        .INPUT_xSyncroPhotocell_1   // M403.P115B1.Synchro photocell / start count
        .PH_x.0   // Load
        .PH_x.1   // Load Upstream
        .PH_x.10   // Unload Upstream
        .PH_x.11   // End load Downstream
        .PH_x.12   // Unload Downstream
        .PH_x.13   // End unload Upstream
        .PH_x.14   // End unload Downstream
        .PH_x.15   // End unload
        .PH_x.16   // Unload Unpack (n caps)
        .PH_x.17   // End unload Unpack (n caps)
        .PH_x.18   // Unload Unpack (n caps) Upstream
        .PH_x.19   // End unload Unpack (n caps) Upstream
        .PH_x.2   // Load Downstream
        .PH_x.20   // Unload Unpack (n caps) Downstream
        .PH_x.21   // End unload Unpack (n caps) Downstream
        .PH_x.22   // Load reentry
        .PH_x.23   // End load reentry
        .PH_x.24   // Unload reentry
        .PH_x.25   // End unload reentry
        .PH_x.26   // Load Unpack (n caps)
        .PH_x.27   // End load Unpack (n caps)
        .PH_x.28   // Load Unpack (n caps) Upstream
        .PH_x.29   // End load Unpack (n caps) Upstream
        .PH_x.3   // Wait rotation done
        .PH_x.30   // Load Unpack (n caps) Downstream
        .PH_x.31   // End load Unpack (n caps) Downstream
        .PH_x.4   // Rotation ended
        .PH_x.7   // End load
        .PH_x.8   // Unload
        .PH_x.9   // End load Upstream
   M316_ALM : MAC_Conveyor_ALM;
        .rgdFaultCode_M[0]   // Drive fault code M1
        .rgdFaultCode_M[1]   // Drive fault code M2
        .rgxStoppingFault[0].0   // Z402.M316-M1.Positioning error
        .rgxStoppingFault[0].1   // Z402.M316-M1.Phase in progress with rotator not in low position
        .rgxStoppingFault_M[0].0   // Z402.M316-M1.Protection motor rotation
        .rgxStoppingFault_M[0].1   // Z402.M316-M1.Drive error
        .rgxStoppingFault_M[0].2   // Z402.M316-M1.Drive feedback error
        .rgxStoppingFault_M[0].3   // Z402.M316-M1.Local safety switch
        .rgxStoppingFault_M[0].4   // Z402.M316-M1.Motor thermal probe
        .rgxStoppingFault_M[0].5   // Z402.M316-M1.Braking resistor anomaly
        .rgxStoppingFault_M[0].6   // Z402.M316-M1.Drive not ready
        .rgxWarning[0].0   // Z402.M316.Plate not synchronized
        .rgxWarning[0].1   // Z402.M316.Positioning error
   M316_Data : UDT_Convoy_SL;
   M316_dLastRotationA_ID : DINT; {access Read Only}
   M316_HMR : MAC_Conveyor_HMR := (xIdPlatePresence := 1, dState1 := 1, dState2 := 1, dStateSensor1 := 1, dStateSensor2 := 1, dStateSensor3 := 1, dStateSensor4 := 1);
        .dErrorCode1   // Error code M1
        .rgxMan.0   // Run M1
        .rgxMan.1   // Reverse M1
        .rgxMan.2   // Run M2
        .rgxMan.3   // Reverse M2
        .rgxMan.4   // Run both
        .rgxMan.5   // Reverse both
        .dErrorCode2   // Error code M2
        .xSensorPresence1   // M403.P115B1.Synchro photocell / start count {x|x|x|x|O}
        .xSensorPresence2   // M403.P115B2.Synchro photocell / start count {x|x|x|x|O}
   M316_HMW : MAC_Conveyor_HMW;
        .dParam_1_cmm   // Positioning offset 1 [mm] {mm/100|mm|-50|+50|M}
        .dParam_2_cmm   // Positioning offset 2 [mm] {mm/100|mm|-50|+50|M}
        .rgxMan.0   // Run M1
        .rgxMan.1   // Reverse M1
        .rgxMan.2   // Run M2
        .rgxMan.3   // Reverse M2
        .rgxMan.4   // Run both
        .rgxMan.5   // Reverse both
   M316_M1_DR : AXIS_CIP_DRIVE; {access Read Only}
   M316_M1_DR_IN_MAJ : MOTION_INSTRUCTION := (FLAGS := 570425344, DN := 1); {access None}
   M316_M1_DR_IN_MAM : MOTION_INSTRUCTION := (FLAGS := 704643072, DN := 1, PC := 1); {access None}
   M316_M1_DR_IN_MAR : MOTION_INSTRUCTION := (FLAGS := 167772160, PC := 1); {access None}
   M316_M1_DR_IN_MAS : MOTION_INSTRUCTION := (FLAGS := -1442840576, EN := 1, DN := 1, PC := 1); {access None}
   M316_M1_DR_IN_MCD : MOTION_INSTRUCTION := (FLAGS := 570425344, DN := 1); {access None}
   M316_M1_DR_IN_MRP : MOTION_INSTRUCTION := (FLAGS := 536870912, DN := 1, STATUS := 2, STATE := 3); {access None}
   M316_M1_DR_MAFR : MOTION_INSTRUCTION := (FLAGS := 301989888, ER := 1, ERR := 11); {access None}
   M316_M1_DR_MDR : MOTION_INSTRUCTION := (FLAGS := -1845493760, EN := 1, ER := 1, ERR := 11); {access None}
   M316_M1_DR_MSF : MOTION_INSTRUCTION := (FLAGS := 570425344, DN := 1, STATUS := 2, STATE := 1); {access None}
   M316_M1_DR_MSO : MOTION_INSTRUCTION := (FLAGS := -1610612736, EN := 1, DN := 1, STATE := 1); {access None}
   M316_M1_DR_OUT_MAJ : MOTION_INSTRUCTION := (FLAGS := 570425344, DN := 1); {access None}
   M316_M1_DR_OUT_MAM : MOTION_INSTRUCTION := (FLAGS := 704643072, DN := 1, PC := 1); {access None}
   M316_M1_DR_OUT_MAR : MOTION_INSTRUCTION := (FLAGS := 671088640, DN := 1, PC := 1, STATE := 1); {access None}
   M316_M1_DR_OUT_MAS : MOTION_INSTRUCTION := (FLAGS := -1442840576, EN := 1, DN := 1, PC := 1); {access None}
   M316_M1_DR_OUT_MCD : MOTION_INSTRUCTION := (FLAGS := 570425344, DN := 1); {access None}
   M316_M1_DR_OUT_MRP : MOTION_INSTRUCTION := (FLAGS := 536870912, DN := 1, STATUS := 2, STATE := 3); {access None}
   M316_SpaceConv_Utilities : SpaceConv_Utilities := (CONST_dSyncMode := 1, CONST_dSyncroPhWindow_cmm := 450000, CONST_dConveyorLength_cmm := 800000, CONST_dConveyorWidth_cmm := 400000, CONST_dPresetFeedbackTime_ms := 500, CONST_rAcceleration_ms2 := 1.2, CONST_rDeceleration_ms2 := 1.2, CONF_MD1_dScan_ms := 20, CONF_MD2_MD3_dPrstPos_cmm := -390000, CONF_MD4_MD6_dLength_cmm := 365800, CONF_MD7_dOffset_cmm := 50000, ST_dStopLoadForseen_cmm := 620000, ST_dRealSpeed_mm_min := 90000, ST_rStepAdvancementH := 3000.0, ST_rStepAdvancementT := 3000.0, O_xPlateSynchronized := 1, O_dCountFeedbackTime_ms := 500, O_dPresetLoadUnload_cmm := -126300);
   M316_TON_Synchro_timeout : TIMER; {access Read Only}
   M316_xOS_SentToCullet : BOOL; {access Read Only}
   M316_xPlateCullet : BOOL; {access Read Only}
   M316_xSendCulletReqActive : BOOL; {access Read Only}
   M316_xSensorTimeout : BOOL; {access Read Only}
   M316A : MAC_Rotator := (ST_xCleaningConditionOK := 1, ST_xConditionOKStopCycle := 1, ST_xEnableControlError := 1, INPUT_rRotatorPosition_cdeg := 26999.898, INPUT_xConditionToDescent := 1, INPUT_xLowPosition := 1, INPUT_xLocalSafetySwitchRotation := 1, INPUT_xProtectionMotorLifting := 1, INPUT_xProtectionMotorRotation := 1, tmON_DelayFrameUP.PRE := 100, tmON_DelayRotatorInRun.PRE := 300, tmOF_DriveEnable.PRE := 20000, tmOF_DriveEnable.ACC := 20000, tmON_FeedbackTimeOutLifting.PRE := 1000, tmON_FeedbackTimeOutRotation.PRE := 1000, tmON_FramePosError.PRE := 2500, tmON_RotatePosError.PRE := 10000, tmON_RotatePosError.ACC := 2040, tmON_RotatePosError.EN := 1, tmON_RotatePosError.TT := 1, tmON_PresetEncoder.PRE := 3000, tmON_DelayBrakeON.PRE := 200); {access None}
        .OUTPUT_xDescent   // P253KA4.Descent frame
        .PH_x.0   // Rise frame
        .PH_x.12   // Counterclockwise rotation
        .PH_x.4   // Descent frame
        .PH_x.8   // Clockwise totation
        .OUTPUT_xRise   // P253KA3.Lifting frame
        .INPUT_xLowPosition   // P56KA2.Frame to low position
        .INPUT_xFeedbackLifting   // P56KM1/2.Feedback lifting chassis
        .INPUT_xHighPosition   // P56KA1.Frame to high position
        .INPUT_xProtectionMotorLifting   // P56QM1.Protection lifting frame
   M316A_ALM : MAC_Rotator_ALM;
        .rgxStoppingFault_M[0].0   // Z402.M316A.Protection motor rotation
        .rgxStoppingFault_M[0].1   // Z402.M316A.Drive Error
        .rgxStoppingFault_M[0].11   // Z402.M316A.Frame lifting position error
        .rgxStoppingFault_M[0].2   // Z402.M316A.Drive feedback error
        .rgxStoppingFault_M[0].20   // Z402.M316A.Drive not ready
        .rgxStoppingFault_M[0].3   // Z402.M316A.Rotation position error
        .rgxStoppingFault_M[0].8   // Z402.M316A.Protection lifting frame
        .rgxStoppingFault_M[0].9   // Z402.M316A.Feedback lifting chassis
   M316A_Data : UDT_Convoy_SL;
   M316A_HMR : MAC_Rotator_HMR := (xLowPosition := 1, dState := 1, dActualAngle_cdeg := 27000);
        .rgxMan.0   // Rise
        .rgxMan.1   // Descent
        .rgxMan.10   // Clockwise rotation jog
        .rgxMan.11   // Counter Clockwise rotation jog
        .rgxMan.14   // Enable brake release
        .rgxMan.15   // Disable brake release
        .rgxMan.8   // Clockwise rotation
        .rgxMan.9   // Counter Clockwise rotation
   M316A_HMW : MAC_Rotator_HMW := (xPresetEnc := 1, dLowSpeed_deg_s := 40, dLowRamp_deg_s2 := 50, dHighSpeed_deg_s := 50, dHighRamp_deg_s2 := 60, dJogSpeed_deg_s := 12);
        .rgxMan.0   // Rise
        .rgxMan.1   // Descent
        .rgxMan.10   // Clockwise rotation jog
        .rgxMan.11   // Counterclockwise rotation jog
        .rgxMan.14   // Enable brake release
        .rgxMan.15   // Disable brake release
        .rgxMan.8   // Clockwise rotation
        .rgxMan.9   // Counterclockwise rotation
   M316A_M1_DR : AXIS_CIP_DRIVE; {access Read Only}
   M316A_M1_DR_IN_MAJ : MOTION_INSTRUCTION := (FLAGS := 570425344, DN := 1); {access None}
   M316A_M1_DR_IN_MAM : MOTION_INSTRUCTION := (FLAGS := 704643072, DN := 1, PC := 1); {access None}
   M316A_M1_DR_IN_MAS : MOTION_INSTRUCTION := (FLAGS := -1442840576, EN := 1, DN := 1, PC := 1); {access None}
   M316A_M1_DR_MAFR : MOTION_INSTRUCTION := (FLAGS := 301989888, ER := 1, ERR := 11); {access None}
   M316A_M1_DR_MAH : MOTION_INSTRUCTION := (FLAGS := 671088640, DN := 1, PC := 1, STATE := 17); {access None}
   M316A_M1_DR_MSF : MOTION_INSTRUCTION := (FLAGS := -1610612736, EN := 1, DN := 1, STATUS := 2, STATE := 1); {access None}
   M316A_M1_DR_MSO : MOTION_INSTRUCTION := (FLAGS := 536870912, DN := 1, STATE := 1); {access None}
   M316A_M1_DR_OUT_MAJ : MOTION_INSTRUCTION := (FLAGS := 570425344, DN := 1); {access None}
   M316A_M1_DR_OUT_MAM : MOTION_INSTRUCTION := (FLAGS := 704643072, DN := 1, PC := 1); {access None}
   M316A_M1_DR_OUT_MAS : MOTION_INSTRUCTION := (FLAGS := -1442840576, EN := 1, DN := 1, PC := 1); {access None}
   M316A_MAM_IP_TOFF : TIMER; {access Read Only}
   M316A_rLastPosition : REAL; {access Read Only}
   M316A_TmON1 : TIMER; {access Read Only}
   M316M317_OffsetBaricentre_cmm : DINT; {access Read Only}
   M317 : MAC_Conveyor_Single := (ST_xCleaningConditionOK := 1, ST_xPlatePresence := 1, ST_xConditionOKStopCycle := 1, ST_xOutputEnable := 1, ST_xIdPlatePresence := 1, ST_xWaitStopNextMachine := 1, ST_xEnableControlError := 1, ST_xPlateSynchronized := 1, ST_xSafetyMovement := 1, OSR_xSynchroPhotocellTail := 1, INPUT_xSquaringPhotocell_4 := 1, INPUT_xLowPositionSquaring_1 := 1, INPUT_xHighPositionPopup_1 := 1, INPUT_xHighPositionPopup_2 := 1, INPUT_xDriveReady_M1 := 1, INPUT_xLocalSafetySwitch_M1 := 1, INPUT_xMotorThermalProbe_M1 := 1, INPUT_xProtectionMotor_M1 := 1, INPUT_xDriveReady_M2 := 1, INPUT_xLocalSafetySwitch_M2 := 1, INPUT_xMotorThermalProbe_M2 := 1, INPUT_xProtectionMotor_M2 := 1, INPUT_xDriveFeedback_M3 := 1, INPUT_xDriveReady_M3 := 1, INPUT_xLocalSafetySwitch_M3 := 1, INPUT_xMotorThermalProbe_M3 := 1, INPUT_xProtectionMotor_M3 := 1, INPUT_xDriveReady_M4 := 1, INPUT_xLocalSafetySwitch_M4 := 1, INPUT_xMotorThermalProbe_M4 := 1, INPUT_xProtectionMotor_M4 := 1, INPUT_xProtectionLiftingFrame_1 := 1, INPUT_xProtectionLiftingFrame_2 := 1, INPUT_xFeedbackVentilation_1 := 1, INPUT_xFeedbackVentilation_2 := 1, OUTPUT_xDriveEnable_M1 := 1, OUTPUT_xDriveEnable_M2 := 1, OUTPUT_xDriveEnable_M3 := 1, OUTPUT_xDriveEnable_M4 := 1, OUTPUT_xFunCommand_1 := 1, OUTPUT_xFunCommand_2 := 1, AUX_dPresetStopLoad_cmm := 372333, AUX_dPresetStopUnload_cmm := 441667, AUX_dAccSpace_cmm := 41667, AUX_dDecSpace_cmm := 41667, AUX_dReqSpeed_mm_min := 60000, AUX_dAbsPosTarget_M3_cmm := 195500, AUX_dAbsPosTarget_M4_cmm := 195500, AUX_dQtaLites := 1, tmON_FeedbackTimeOut_M1.PRE := 2000, tmOF_DriveEnable_M1.PRE := 30000, tmOF_DriveEnable_M1.ACC := 540, tmOF_DriveEnable_M1.TT := 1, tmOF_DriveEnable_M1.DN := 1, tmOF_PowerSaving_M1.EN := 1, tmOF_PowerSaving_M1.DN := 1, tmON_FeedbackTimeOut_M2.PRE := 2000, tmOF_DriveEnable_M2.PRE := 30000, tmOF_DriveEnable_M2.ACC := 540, tmOF_DriveEnable_M2.TT := 1,
        tmOF_DriveEnable_M2.DN := 1, tmON_FeedbackTimeOut_M3.PRE := 2000, tmOF_DriveEnable_M3.PRE := 30000, tmOF_DriveEnable_M3.ACC := 540, tmOF_DriveEnable_M3.TT := 1, tmOF_DriveEnable_M3.DN := 1, tmON_FeedbackTimeOut_M4.PRE := 2000, tmOF_DriveEnable_M4.PRE := 30000, tmOF_DriveEnable_M4.ACC := 540, tmOF_DriveEnable_M4.TT := 1, tmOF_DriveEnable_M4.DN := 1, tmON_AuxFunction1.PRE := 5000, tmON_AuxFunction1.EN := 1, tmON_AuxFunction1.DN := 1, tmON_AuxFunction2.PRE := 2200, tmON_AuxFunction3.PRE := 2200, tmON_AuxFunction4.PRE := 15000, tmON_AuxFunction5.PRE := 3000, tmON_AuxFunction6.PRE := 15000, tmON_AuxFunction7.PRE := 3600000, tmON_AuxFunction8.PRE := 40000, tmON_AuxFunction9.PRE := 20000, TmON[0].PRE := 3000, TmON[1].PRE := 1000, TmON[1].ACC := 1019, TmON[2].PRE := 5000, TmON[6].PRE := 5000, TmON[6].EN := 1, TmON[6].DN := 1, TmON[11].PRE := 2000, TmON[12].PRE := 2000, TmON[13].PRE := 2000, TmON[14].PRE := 2000, tmOF_MCD_M1.ACC := 20, tmOF_MCD_M2.ACC := 20, tmOF_MCD_M3.ACC := 20, tmOF_MCD_M4.ACC := 20); {access None}
        .INPUT_xSquaringPhotocell_1   // P406B1.Squaring frontal photocell - Right
        .INPUT_xMotorThermalProbe_M2   // M2.P404BT2.Motor thermal probe
        .INPUT_xLowPositionPopup_1   // P63KA2.M5.Low position popup
        .INPUT_xLowPositionSquaring_1   // P405SQ2.Low position squaring
        .INPUT_xMotorThermalProbe_M1   // M1.P404BT1.Motor thermal probe
        .INPUT_xHighPositionPopup_1   // P63KA1.M5.High position popup
        .INPUT_xSquaringPhotocell_2   // P406B2.Squaring frontal photocell - Left
        .INPUT_xHighPositionPopup_2   // P64KA1.M6.High position popup
        .PH_x.0   // Load (from M316)
        .PH_x.10   // Load (from M419)
        .PH_x.11   // End load (from M419)
        .PH_x.12   // Unload (to M316)
        .PH_x.13   // End unload (to M316)
        .PH_x.15   // End unload (to M419)
        .PH_x.16   // Rise popup
        .PH_x.19   // End rise popup
        .PH_x.20   // Descent popup
        .PH_x.23   // End descent popup
        .PH_x.24   // Reset counter position
        .PH_x.26   // Lateral positioning (M3-M4)
        .PH_x.27   // End lateral positioning (M3-M4)
        .PH_x.28   // Lateral squaring
        .PH_x.29   // End lateral squaring
        .PH_x.30   // Lateral traction recovery (M3-M4)
        .PH_x.31   // End lateral traction recovery (M3-M4)
        .PH_x.4   // Frontal squaring (run fwd + rise squaring)
        .PH_x.5   // End frontal sqauring
        .PH_x.7   // End load (from M316)
        .PH_x.8   // Unload (to M419)
        .INPUT_xMotorThermalProbe_M3   // M3.P405BT3.Motor thermal probe
        .INPUT_xLowPositionPopup_2   // P64KA2.M6.Low position popup
        .INPUT_xSquaringPhotocell_3   // P405B1.Squaring lateral photocell - Right
        .INPUT_xHighPositionSquaring_1   // P405SQ1.High position squaring
        .INPUT_xSquaringPhotocell_4   // P405B2.Squaring lateral photocell - Left
        .INPUT_xHighPositionSquaring_2   // P405SQ11.High position squaring
        .ST_xAux1   // Ready to unload on backward conveyor
        .INPUT_xLowPositionSquaring_2   // P405SQ12.Low position squaring
   M317_ALM : MAC_Conveyor_ALM;
        .rgxWarning[0].10   // Z402.M317-M2.Plate not synchronized
        .rgdFaultCode_M[0]   // Drive fault code M1
        .rgdFaultCode_M[1]   // Drive fault code M2
        .rgxStoppingFault[0].0   // Z402.M317-M1.Positioning error
        .rgxStoppingFault[0].1   // Z402.M317-M1.Plate not synchronized
        .rgxStoppingFault[0].10   // Z402.M317-M2.Error position frontal squaring
        .rgxStoppingFault[0].11   // Z402.M317-M2.Timeout frontal squaring
        .rgxStoppingFault[0].12   // Z402.M317-M2.Lugs position sensors fault
        .rgxStoppingFault[0].13   // Z402.M317. Timeout movement popup 1
        .rgxStoppingFault[0].14   // Z402.M317. Timeout movement popup 2
        .rgxStoppingFault[0].16   // Z402.M317-M3.Positioning error
        .rgxStoppingFault[0].18   // Z402.M317-M3.Error position popup
        .rgxStoppingFault[0].19   // Z402.M317-M3.Error position lateral squaring
        .rgxStoppingFault[0].2   // Z402.M317-M1.Error position frontal squaring
        .rgxStoppingFault[0].20   // Z402.M317-M3.Timeout lateral squaring
        .rgxStoppingFault[0].21   // Z402.M317.Protection lifting popup 1
        .rgxStoppingFault[0].22   // Z402.M317.Protection lifting popup 2
        .rgxStoppingFault[0].3   // Z402.M317-M1.Timeout frontal squaring
        .rgxStoppingFault[0].4   // Z402.M317-M1.Lugs position sensors fault
        .rgxStoppingFault[0].5   // Z402.M317. Popup 1 position error
        .rgxStoppingFault[0].6   // Z402.M317. Popup 2 position error
        .rgxStoppingFault[0].8   // Z402.M317-M2.Positioning error
        .rgxStoppingFault[0].9   // Z402.M317-M2.Plate not synchronized
        .rgxStoppingFault_M[0].0   // Z402.M317-M1.P59AZ1.Protection motor rotation
        .rgxStoppingFault_M[0].1   // Z402.M317-M1.P59AZ1.Drive error
        .rgxStoppingFault_M[0].10   // Z402.M317-M2.P59AZ1.Drive feedback error
        .rgxStoppingFault_M[0].11   // Z402.M317-M2.P59AZ1.Local safety switch
        .rgxStoppingFault_M[0].12   // Z402.M317-M2.P405BT2.Motor thermal probe
        .rgxStoppingFault_M[0].13   // Z402.M317-M2.P59AZ1.Braking resistor anomaly
        .rgxStoppingFault_M[0].14   // Z402.M317-M2.Drive not ready
        .rgxStoppingFault_M[0].16   // Z402.M317-M3.P61AZ1.Protection motor rotation
        .rgxStoppingFault_M[0].17   // Z402.M317-M3.P61AZ1.Drive error
        .rgxStoppingFault_M[0].18   // Z402.M317-M3.P61AZ1.Drive feedback error
        .rgxStoppingFault_M[0].19   // Z402.M317-M3.P61AZ1.Local safety switch
        .rgxStoppingFault_M[0].2   // Z402.M317-M1.P59AZ1.Drive feedback error
        .rgxStoppingFault_M[0].20   // Z402.M317-M3.P404BT1.Motor thermal probe
        .rgxStoppingFault_M[0].21   // Z402.M317-M3.Drive not ready
        .rgxStoppingFault_M[0].3   // Z402.M317-M1.P59AZ1.Local safety switch
        .rgxStoppingFault_M[0].4   // Z402.M317-M1.P405BT1.Motor thermal probe
        .rgxStoppingFault_M[0].5   // Z402.M317-M1.P59AZ1.Braking resistor anomaly
        .rgxStoppingFault_M[0].6   // Z402.M317-M1.Drive not ready
        .rgxStoppingFault_M[0].8   // Z402.M317-M2.P59AZ1.Protection motor rotation
        .rgxStoppingFault_M[0].9   // Z402.M317-M2.P59AZ1.Drive error
        .rgxWarning[0].0   // Z402.M317-M1.Plate not synchronized
        .rgxWarning[0].1   // Z402.M317-M1.Positioning error
        .rgxWarning[0].11   // Z402.M317-M2.Positioning error
        .rgxWarning[0].21   // Z402.M317-M3.Lateal positioning error
        .rgxWarning[0].25   // Z402.M317.Timeout frontal squaring
        .rgxWarning[0].26   // Z402.M317.Timeout lateral squaring
   M317_AlmTimer1 : TIMER; {access Read Only}
   M317_AlmTimer2 : TIMER; {access Read Only}
   M317_Data : UDT_Convoy_SL;
        .rgtCap[0].rgxRequest.0   // Frontal squaring request
        .rgtCap[0].rgxRequest.1   // Lateral squaring request
        .rgtCap[0].rgxRequest.2   // Y adjust position request
        .rgtCap[0].rgxRequest.3   // Y measure request
        .rgtCap[0].rgxDone.0   // Frontal squaring done
        .rgtCap[0].rgxDone.1   // Lateral squaring done
        .rgtCap[0].rgxDone.2   // Y adjust position done
        .rgtCap[0].rgxDone.3   // Y measure done
   M317_dSlowingSquaringQuote : DINT; {access Read Only}
   M317_dTractionRecovery_M3 : DINT; {access Read Only}
   M317_dTractionRecovery_M4 : DINT; {access Read Only}
   M317_HMR : MAC_Conveyor_HMR := (xSensorPresence4 := 1, xHighPositionPopup1 := 1, xHighPositionPopup2 := 1, xLowPositionSquaring1 := 1, xLowPositionSquaring2 := 1, xIdPlatePresence := 1, dState1 := 1, dState2 := 1, dState3 := 1, dState4 := 1, dStateSensor1 := 1, dStateSensor2 := 1, dStateSensor3 := 1, dStateSensor4 := 1, dStateSensor5 := 1, dStateSensor6 := 1);
        .xSensorPresence5   // P115/3.Start count photocell {x|x|x|x|O}
        .xHighPositionPopup2   // P64KA1.M6.High position popup {x|x|x|x|O}
        .dErrorCode1   // Error code M1
        .xHighPositionPopup1   // P63KA1.M5.High position popup {x|x|x|x|O}
        .rgxMan.0   // Run M1
        .rgxMan.1   // Reverse M1
        .rgxMan.10   // Rise popup 1
        .rgxMan.11   // Descent popup 1
        .rgxMan.12   // Rise popup 2
        .rgxMan.13   // Descent popup 2
        .rgxMan.14   // Rise all popups
        .rgxMan.15   // Descent all popups
        .rgxMan.16   // Rise frontal squaring 1
        .rgxMan.17   // Descent frontal squaring 1
        .rgxMan.18   // Rise frontal squaring 2
        .rgxMan.19   // Descent frontal squaring 2
        .rgxMan.2   // Run M2
        .rgxMan.20   // Rise all frontal squaring
        .rgxMan.21   // Descent all frontal squaring
        .rgxMan.3   // Reverse M2
        .rgxMan.4   // Run M3
        .rgxMan.5   // Reverse M3
        .rgxMan.6   // Run M4
        .rgxMan.7   // Reverse M4
        .dState3   // State M3 (1=No anomaly; 3=Run; 4=Reverse; 7=Anomaly)
        .xHighPositionSquaring1   // P405SQ1.High position frontal squaring M1 {x|x|x|x|O}
        .dErrorCode2   // Error code M2
        .xSensorPresence6   // P115/4.Start count photocell {x|x|x|x|O}
        .xSensorPresence4   // P404B1.SlowDown photocell frontal squaring left {x|x|x|x|O}
        .xLowPositionPopup1   // P63KA2.M5.Low position popup {x|x|x|x|O}
        .xHighPositionSquaring2   // P405SQ11.High position frontal squaring M2 {x|x|x|x|O}
        .dState2   // State M2 (1=No anomaly; 3=Run; 4=Reverse; 7=Anomaly)
        .dErrorCode4   // Error code M4
        .xSensorPresence3   // P404B1.SlowDown photocell frontal squaring right {x|x|x|x|O}
        .dState1   // State M1 (1=No anomaly; 3=Run; 4=Reverse; 7=Anomaly)
        .dState4   // State M4 (1=No anomaly; 3=Run; 4=Reverse; 7=Anomaly)
        .xLowPositionSquaring2   // P405SQ12.Low position frontal squaring M2 {x|x|x|x|O}
        .xLowPositionSquaring1   // P405SQ2.Low position frontal squaring M1 {x|x|x|x|O}
        .xLowPositionPopup2   // P64KA2.M6.Low position popup {x|x|x|x|O}
        .xSensorPresence1   // P405B1.SlowDown photocell lateral squaring right {x|x|x|x|O}
        .dErrorCode3   // Error code M3
        .xSensorPresence2   // P405B2.SlowDown photocell lateral squaring left {x|x|x|x|O}
   M317_HMW : MAC_Conveyor_HMW := (dParam_3_cmm := 4000, dParam_5_ms := 3000, dParam_6_ms := 4000, dParam_7_ms := 2200, dParam_8_ms := 5000);
        .dParam_4_cmm   // Lateral squaring space {mm/100|mm|0|500|M}
        .dParam_1_cmm   // Positioning offset 1 {mm/100|mm|-50|+50|M}
        .dParam_3_cmm   // Frontal squaring space {mm/100|mm|0|500|M}
        .dParam_6_ms   // Squaring frontal time 2 {ms|s|0|5|M}
        .dParam_2_cmm   // Positioning offset 2 {mm/100|mm|-50|+50|M}
        .dParam_8_ms   // Squaring lateral time 2 {ms|s|0|5|M}
        .rgxMan.0   // Run M1
        .rgxMan.1   // Reverse M1
        .rgxMan.10   // Rise popup 2
        .rgxMan.11   // Descent popup 2
        .rgxMan.12   // Rise all popups
        .rgxMan.13   // Descent all popups
        .rgxMan.14   // Run both (M1-2)
        .rgxMan.15   // Reverse both (M1-2)
        .rgxMan.16   // Rise frontal squaring 1
        .rgxMan.17   // Descent frontal squaring 1
        .rgxMan.18   // Rise frontal squaring 2
        .rgxMan.19   // Descent frontal squaring 2
        .rgxMan.2   // Run M2
        .rgxMan.20   // Rise all frontal squaring
        .rgxMan.21   // Descent all frontal squaring
        .rgxMan.3   // Reverse M2
        .rgxMan.4   // Run M3
        .rgxMan.5   // Reverse M3
        .rgxMan.6   // Run M4
        .rgxMan.7   // Reverse M4
        .rgxMan.8   // Rise popup 1
        .rgxMan.9   // Descent popup 1
        .dParam_7_ms   // Squaring lateral time 1 {ms|s|0|5|M}
        .dParam_5_ms   // Squaring frontal time 1 {ms|s|0|5|M}
   M317_M1_DR_IN_MAJ : MOTION_INSTRUCTION := (FLAGS := 570425344, DN := 1); {access None}
   M317_M1_DR_IN_MAM : MOTION_INSTRUCTION := (FLAGS := 33554432); {access None}
   M317_M1_DR_IN_MAR : MOTION_INSTRUCTION := (FLAGS := 33554432); {access None}
   M317_M1_DR_IN_MAS : MOTION_INSTRUCTION := (FLAGS := -1442840576, EN := 1, DN := 1, PC := 1); {access None}
   M317_M1_DR_IN_MCD : MOTION_INSTRUCTION := (FLAGS := 570425344, DN := 1); {access None}
   M317_M1_DR_IN_MRP : MOTION_INSTRUCTION := (FLAGS := 33554432); {access None}
   M317_M1_DR_MAFR : MOTION_INSTRUCTION := (FLAGS := 301989888, ER := 1, ERR := 11); {access None}
   M317_M1_DR_MDR : MOTION_INSTRUCTION := (FLAGS := -1845493760, EN := 1, ER := 1, ERR := 11); {access None}
   M317_M1_DR_MSF : MOTION_INSTRUCTION := (FLAGS := 570425344, DN := 1, STATUS := 2, STATE := 1); {access None}
   M317_M1_DR_MSO : MOTION_INSTRUCTION := (FLAGS := -1610612736, EN := 1, DN := 1, STATE := 1); {access None}
   M317_M1_DR_OUT_MAJ : MOTION_INSTRUCTION := (FLAGS := 570425344, DN := 1); {access None}
   M317_M1_DR_OUT_MAM : MOTION_INSTRUCTION := (FLAGS := 33554432); {access None}
   M317_M1_DR_OUT_MAR : MOTION_INSTRUCTION := (FLAGS := 33554432); {access None}
   M317_M1_DR_OUT_MAS : MOTION_INSTRUCTION := (FLAGS := -1442840576, EN := 1, DN := 1, PC := 1); {access None}
   M317_M1_DR_OUT_MCD : MOTION_INSTRUCTION := (FLAGS := 570425344, DN := 1); {access None}
   M317_M1_DR_OUT_MRP : MOTION_INSTRUCTION := (FLAGS := 33554432); {access None}
   M317_M1_DR_R1 : AXIS_CIP_DRIVE; {access Read Only}
   M317_M2_AUX_ReqSpeed_mm_min : DINT; {access Read Only}
   M317_M2_ChangeSpeed : BOOL; {access Read Only}
   M317_M2_DR_IN_MAJ : MOTION_INSTRUCTION := (FLAGS := 570425344, DN := 1); {access None}
   M317_M2_DR_IN_MAM : MOTION_INSTRUCTION := (FLAGS := 33554432); {access None}
   M317_M2_DR_IN_MAR : MOTION_INSTRUCTION := (FLAGS := 33554432); {access None}
   M317_M2_DR_IN_MAS : MOTION_INSTRUCTION := (FLAGS := 704643072, DN := 1, PC := 1); {access None}
   M317_M2_DR_IN_MCD : MOTION_INSTRUCTION := (FLAGS := 301989888, ER := 1, ERR := 23); {access None}
   M317_M2_DR_IN_MRP : MOTION_INSTRUCTION := (FLAGS := 536870912, DN := 1, STATUS := 2, STATE := 3); {access None}
   M317_M2_DR_MAFR : MOTION_INSTRUCTION := (FLAGS := 301989888, ER := 1, ERR := 11); {access None}
   M317_M2_DR_MDR : MOTION_INSTRUCTION := (FLAGS := -1845493760, EN := 1, ER := 1, ERR := 11); {access None}
   M317_M2_DR_MSF : MOTION_INSTRUCTION := (FLAGS := 570425344, DN := 1, STATUS := 2, STATE := 1); {access None}
   M317_M2_DR_MSO : MOTION_INSTRUCTION := (FLAGS := -1610612736, EN := 1, DN := 1, STATE := 1); {access None}
   M317_M2_DR_OUT_MAJ : MOTION_INSTRUCTION := (FLAGS := 570425344, DN := 1); {access None}
   M317_M2_DR_OUT_MAM : MOTION_INSTRUCTION := (FLAGS := 33554432); {access None}
   M317_M2_DR_OUT_MAR : MOTION_INSTRUCTION := (FLAGS := 33554432); {access None}
   M317_M2_DR_OUT_MAS : MOTION_INSTRUCTION := (FLAGS := 704643072, DN := 1, PC := 1); {access None}
   M317_M2_DR_OUT_MCD : MOTION_INSTRUCTION := (FLAGS := 301989888, ER := 1, ERR := 23); {access None}
   M317_M2_DR_OUT_MRP : MOTION_INSTRUCTION := (FLAGS := 536870912, DN := 1, STATUS := 2, STATE := 3); {access None}
   M317_M2_DR_R2 : AXIS_CIP_DRIVE; {access Read Only}
   M317_M2_ReqSpeed_mm_min : DINT; {access Read Only}
   M317_M3_AUX_ReqSpeed_mm_min : DINT; {access Read Only}
   M317_M3_ChangeSpeed : BOOL; {access Read Only}
   M317_M3_DR_IN_MAJ : MOTION_INSTRUCTION := (FLAGS := 570425344, DN := 1); {access None}
   M317_M3_DR_IN_MAM : MOTION_INSTRUCTION := (FLAGS := -1509949440, EN := 1, DN := 1, IP := 1); {access None}
   M317_M3_DR_IN_MAR : MOTION_INSTRUCTION := (FLAGS := 33554432); {access None}
   M317_M3_DR_IN_MAS : MOTION_INSTRUCTION := (FLAGS := 704643072, DN := 1, PC := 1); {access None}
   M317_M3_DR_IN_MCD : MOTION_INSTRUCTION := (FLAGS := 570425344, DN := 1); {access None}
   M317_M3_DR_IN_MRP : MOTION_INSTRUCTION := (FLAGS := 536870912, DN := 1, STATUS := 2, STATE := 3); {access None}
   M317_M3_DR_L : AXIS_CIP_DRIVE; {access Read Only}
   M317_M3_DR_MAFR : MOTION_INSTRUCTION := (FLAGS := 301989888, ER := 1, ERR := 11); {access None}
   M317_M3_DR_MDR : MOTION_INSTRUCTION := (FLAGS := -1845493760, EN := 1, ER := 1, ERR := 11); {access None}
   M317_M3_DR_MSF : MOTION_INSTRUCTION := (FLAGS := 570425344, DN := 1, STATUS := 2, STATE := 1); {access None}
   M317_M3_DR_MSO : MOTION_INSTRUCTION := (FLAGS := -1610612736, EN := 1, DN := 1, STATE := 1); {access None}
   M317_M3_DR_OUT_MAJ : MOTION_INSTRUCTION := (FLAGS := 570425344, DN := 1); {access None}
   M317_M3_DR_OUT_MAM : MOTION_INSTRUCTION := (FLAGS := -1509949440, EN := 1, DN := 1, IP := 1);
   M317_M3_DR_OUT_MAR : MOTION_INSTRUCTION := (FLAGS := 33554432); {access None}
   M317_M3_DR_OUT_MAS : MOTION_INSTRUCTION := (FLAGS := 704643072, DN := 1, PC := 1); {access None}
   M317_M3_DR_OUT_MCD : MOTION_INSTRUCTION := (FLAGS := 570425344, DN := 1); {access None}
   M317_M3_DR_OUT_MRP : MOTION_INSTRUCTION := (FLAGS := 536870912, DN := 1, STATUS := 2, STATE := 3); {access None}
   M317_M3_ReqSpeed_mm_min : DINT; {access Read Only}
   M317_M3_xOSR_LatSquarFtc : BOOL; {access Read Only}
   M317_SpaceConv_Utilities : SpaceConv_Utilities := (CONST_dSyncMode := 1, CONST_dSyncroPhWindow_cmm := 450000, CONST_dConveyorLength_cmm := 800000, CONST_dConveyorWidth_cmm := 400000, CONST_dPresetFeedbackTime_ms := 500, CONST_rAcceleration_ms2 := 1.2, CONST_rDeceleration_ms2 := 1.2, CONF_MD1_dScan_ms := 20, CONF_MD2_MD3_dPrstPos_cmm := -390000, CONF_MD4_MD6_dLength_cmm := 365800, CONF_MD7_dOffset_cmm := 50000, ST_dStopLoadForseen_cmm := 620000, ST_dRealSpeed_mm_min := 90000, ST_rStepAdvancementH := 3000.0, ST_rStepAdvancementT := 3000.0, O_xPlateSynchronized := 1, O_dCountFeedbackTime_ms := 500, O_dPresetLoadUnload_cmm := -126300);
   M317_TimerAlm3 : TIMER; {access Read Only}
   M317_TON_FrontSquarLeft_timeout : TIMER; {access Read Only}
   M317_TON_FrontSquarRight_timeout : TIMER; {access Read Only}
   M317_TON_LatSquarLeft_timeout : TIMER; {access Read Only}
   M317_TON_LatSquarRight_timeout : TIMER; {access Read Only}
   M317_TON_Load : TIMER; {access Read Only}
   M317_TON_Synchro_timeout : TIMER; {access Read Only}
   M317_xEnableTractionRecovering : BOOL; {access Read Only}
   M317_xFrontLeftTimeout : BOOL; {access Read Only}
   M317_xFrontRightTimeout : BOOL; {access Read Only}
   M317_xLateralTractionRecovered : BOOL; {access Read Only}
   M317_xLatLeftTimeout : BOOL; {access Read Only}
   M317_xLatRightTimeout : BOOL; {access Read Only}
   M317_xOS_PosReq : BOOL;
   M317_xPlateCullet : BOOL; {access Read Only}
   M317_xSendCulletReqActive : BOOL; {access Read Only}
   M317_xSensorTimeout : BOOL; {access Read Only}
   M350_M1_DR : AXIS_CIP_DRIVE; {access Read Only}
   M350_xReqStopPrevConvForPos : BOOL; {access Read Only}
   M350Popup : MAC_Popup_ZC; {access Read Only}
   M350Popup_ALM : MAC_Popup_ZC_ALM; {access Read Only}
        .rgxStoppingFault[0].0   // M350.Lifting position error
   M350Popup_DATA : UDT_ConvoyCap_ZC; {access Read Only}
   M350Popup_HMR : MAC_Popup_ZC_HMR := (xLowPosition := 1, rgdState := 1); {access Read Only}
        .rgxMan.0   // Rise popup {x|x|x|x|O}
        .rgxMan.1   // Lower popup {x|x|x|x|O}
   M350Popup_HMW : MAC_Popup_ZC_HMW := (dSingleCapOffset_cmm := 30000, dGlassPosFromStart_cmm := 15000, dGlassPosFromEnd_cmm := 15000, dConvoySidePosForCenterSheet := 1, dConvoyGapForCenterSheet := 50000, dSaturationSelection := 3);
        .rgxMan.0   // Rise popup {x|x|x|x|O}
        .rgxMan.1   // Lower popup {x|x|x|x|O}
   M350Popup_IN_MOTION : MAC_Popup_ZC_IN_MOTION; {access None}
   M350Popup_OUT_MOTION : MAC_Popup_ZC_OUT_MOTION; {access None}
   M350Popup_PlateFreeTimeout : TIMER := (PRE := 5000); {access Read Only}
   M350Popup_ReentryCap : UDT_ConvoyCap_ZC;
   M350Popup_SearchResultAfter : GP_TrackingSearchPlate_STC;
   M350Popup_SL_DATA : UDT_Convoy_SL; {access Read Only}
   M350Popup_xDrivePosEnable : BOOL; {access Read Only}
   M350Popup_xQualityComing : BOOL; {access Read Only}
   M351 : MAC_Conveyor;
        .INPUT_xMotorThermalProbe_M1   // M315A.M1.Q403BT3. Motor thermal probe
        .PH_x.0   // Load
        .PH_x.1   // Load Upstream
        .PH_x.10   // Unload Downstream
        .PH_x.13   // End unload Upstream
        .PH_x.14   // End unload Downstream
        .PH_x.15   // End unload
        .PH_x.16   // Unpack convoy
        .PH_x.17   // End unpack convoy
        .PH_x.18   // Unpack convoy Upstream
        .PH_x.19   // End unpack convoy Upstream
        .PH_x.2   // Load Downstream
        .PH_x.20   // Unpack convoy Downstream
        .PH_x.21   // End unpack convoy Downstream
        .PH_x.22   // Stop for unload on main line
        .PH_x.23   // End stop for unload on main line
        .PH_x.24   // Stop for unload on main line Upstream
        .PH_x.25   // End stop for unload on main line Upstream
        .PH_x.26   // Stop for unload on main line Downstream
        .PH_x.27   // End stop for unload on main line Downstream
        .PH_x.28   // Load reentry
        .PH_x.29   // End load reentry
        .PH_x.5   // End load Upstream
        .PH_x.6   // End load Downstream
        .PH_x.7   // End load
        .PH_x.8   // Unload
        .PH_x.9   // Unload Upstream
   M351_ALM : MAC_Conveyor_ALM;
        .rgdFaultCode_M[0]   // Drive fault code
        .rgxStoppingFault_M[0].0   // Z900.M351-M1.Protection motor rotation
        .rgxStoppingFault_M[0].1   // Z900.M351-M1.Drive error
        .rgxStoppingFault_M[0].2   // Z900.M351-M1.Drive feedback error
        .rgxStoppingFault_M[0].3   // Z900.M351-M1.Local safety switch
        .rgxStoppingFault_M[0].4   // Z900.M351.M1. Motor thermal probe
        .rgxStoppingFault_M[0].5   // Z900.M351-M1.Braking resistor anomaly
        .rgxStoppingFault_M[0].6   // Z900.M351-M1.Drive not ready
   M351_Data : UDT_Convoy_SL;
   M351_HMR : MAC_Conveyor_HMR := (xManualCommandEnabled := 1, dState4 := 1);
        .dErrorCode1   // Error code M1
        .rgxMan.0   // Run M1
        .rgxMan.1   // Reverse M1
        .rgxMan.2   // Run M2
        .rgxMan.3   // Reverse M2
        .rgxMan.4   // Run M3
        .rgxMan.5   // Reverse M3
        .dErrorCode2   // Error code M2 (NU)
        .dErrorCode3   // Error code M3 (NU)
   M351_HMW : MAC_Conveyor_HMW;
        .rgxMan.0   // Run M1
        .rgxMan.1   // Reverse M1
        .rgxMan.2   // Run M2
        .rgxMan.3   // Reverse M2
        .rgxMan.4   // Run M3
        .rgxMan.5   // Reverse M3
   M351_M1_DR : AXIS_CIP_DRIVE; {access Read Only}
   M351_M1_DR_IN_MAJ : MOTION_INSTRUCTION := (FLAGS := 570425344, DN := 1); {access None}
   M351_M1_DR_IN_MAM : MOTION_INSTRUCTION := (FLAGS := 33554432); {access None}
   M351_M1_DR_IN_MAR : MOTION_INSTRUCTION := (FLAGS := 33554432); {access None}
   M351_M1_DR_IN_MAS : MOTION_INSTRUCTION := (FLAGS := -1442840576, EN := 1, DN := 1, PC := 1); {access None}
   M351_M1_DR_IN_MCD : MOTION_INSTRUCTION := (FLAGS := 570425344, DN := 1); {access None}
   M351_M1_DR_IN_MRP : MOTION_INSTRUCTION := (FLAGS := 33554432); {access None}
   M351_M1_DR_MAFR : MOTION_INSTRUCTION := (FLAGS := 301989888, ER := 1, ERR := 11); {access None}
   M351_M1_DR_MDR : MOTION_INSTRUCTION := (FLAGS := -1845493760, EN := 1, ER := 1, ERR := 11); {access None}
   M351_M1_DR_MSF : MOTION_INSTRUCTION := (FLAGS := 536870912, DN := 1, STATUS := 2, STATE := 1); {access None}
   M351_M1_DR_MSO : MOTION_INSTRUCTION := (FLAGS := -1577058304, EN := 1, DN := 1, STATE := 1); {access None}
   M351_M1_DR_OUT_MAJ : MOTION_INSTRUCTION := (FLAGS := 570425344, DN := 1); {access None}
   M351_M1_DR_OUT_MAM : MOTION_INSTRUCTION := (FLAGS := 33554432); {access None}
   M351_M1_DR_OUT_MAR : MOTION_INSTRUCTION := (FLAGS := 33554432); {access None}
   M351_M1_DR_OUT_MAS : MOTION_INSTRUCTION := (FLAGS := -1442840576, EN := 1, DN := 1, PC := 1); {access None}
   M351_M1_DR_OUT_MCD : MOTION_INSTRUCTION := (FLAGS := 570425344, DN := 1); {access None}
   M351_M1_DR_OUT_MRP : MOTION_INSTRUCTION := (FLAGS := 33554432); {access None}
   M351_SpaceConv_Utilities : SpaceConv_Utilities := (CONST_dSyncMode := 1, CONST_dSyncroPhWindow_cmm := 200000, CONST_dConveyorLength_cmm := 500000, CONST_dConveyorWidth_cmm := 400000, CONST_dPresetFeedbackTime_ms := 500, CONST_rAcceleration_ms2 := 1.2, CONST_rDeceleration_ms2 := 1.2, CONF_MD1_dScan_ms := 20, CONF_MD4_MD6_dLength_cmm := 360000, CONF_MD7_dOffset_cmm := 50000, ST_xLastModLoadBkw := 1, ST_dStopLoadForseen_cmm := 495370, ST_dRealSpeed_mm_min := 40000, ST_rStepAdvancementH := 1333.3334, ST_rStepAdvancementT := 1333.3334, O_xPlateSynchronized := 1, O_dCountFeedbackTime_ms := 500, O_dPresetLoadUnload_cmm := -440770);
   M352 : MAC_Conveyor;
        .PH_x.25   // End stop for unload on main line Upstream
        .PH_x.0   // Load
        .PH_x.8   // Unload
        .PH_x.24   // Stop for unload on main line Upstream
        .PH_x.21   // End unpack convoy Downstream
        .PH_x.22   // Stop for unload on main line
        .PH_x.23   // End stop for unload on main line
        .PH_x.28   // Load reentry
        .PH_x.29   // End load reentry
        .PH_x.5   // End load Upstream
        .PH_x.6   // End load Downstream
        .PH_x.7   // End load
        .PH_x.9   // Unload Upstream
        .INPUT_xMotorThermalProbe_M1   // M315A.M1.Q403BT3. Motor thermal probe
        .PH_x.1   // Load Upstream
        .PH_x.10   // Unload Downstream
        .PH_x.13   // End unload Upstream
        .PH_x.14   // End unload Downstream
        .PH_x.15   // End unload
        .PH_x.16   // Unpack convoy
        .PH_x.17   // End unpack convoy
        .PH_x.18   // Unpack convoy Upstream
        .PH_x.19   // End unpack convoy Upstream
        .PH_x.2   // Load Downstream
        .PH_x.20   // Unpack convoy Downstream
        .PH_x.26   // Stop for unload on main line Downstream
        .PH_x.27   // End stop for unload on main line Downstream
   M352_ALM : MAC_Conveyor_ALM;
        .rgdFaultCode_M[0]   // Drive fault code
        .rgxStoppingFault_M[0].1   // Z900.M352-M1.Drive error
        .rgxStoppingFault_M[0].6   // Z900.M352-M1.Drive not ready
        .rgxStoppingFault_M[0].0   // Z900.M352-M1.Protection motor rotation
        .rgxStoppingFault_M[0].2   // Z900.M352-M1.Drive feedback error
        .rgxStoppingFault_M[0].3   // Z900.M352-M1.Local safety switch
        .rgxStoppingFault_M[0].4   // Z900.M352.M1. Motor thermal probe
        .rgxStoppingFault_M[0].5   // Z900.M352-M1.Braking resistor anomaly
   M352_Data : UDT_Convoy_SL;
   M352_DeletePlate : BOOL;
   M352_HMR : MAC_Conveyor_HMR := (xManualCommandEnabled := 1, dState4 := 1);
        .rgxMan.0   // Run M1
        .rgxMan.2   // Run M2
        .rgxMan.4   // Run M3
        .dErrorCode1   // Error code M1
        .rgxMan.1   // Reverse M1
        .rgxMan.3   // Reverse M2
        .rgxMan.5   // Reverse M3
        .dErrorCode2   // Error code M2 (NU)
        .dErrorCode3   // Error code M3 (NU)
   M352_HMW : MAC_Conveyor_HMW;
        .rgxMan.0   // Run M1
        .rgxMan.2   // Run M2
        .rgxMan.4   // Run M3
        .rgxMan.1   // Reverse M1
        .rgxMan.3   // Reverse M2
        .rgxMan.5   // Reverse M3
   M352_Input_xPbDeleteGlass : BOOL;
   M352_Input_xPbFanOff : BOOL;   // W204SB3/A. Fan off
   M352_Input_xPbReqGlass : BOOL;   // W204SB1. Request sheet glass
   M352_Input_xPbSendToCullet : BOOL;   // W204SB2. Send to cullet
   M352_INPUT_xSLFanOn : BOOL;
   M352_M1_DR : AXIS_CIP_DRIVE; {access Read Only}
   M352_M1_DR_IN_MAJ : MOTION_INSTRUCTION := (FLAGS := 570425344, DN := 1); {access None}
   M352_M1_DR_IN_MAM : MOTION_INSTRUCTION := (FLAGS := 33554432); {access None}
   M352_M1_DR_IN_MAR : MOTION_INSTRUCTION := (FLAGS := 33554432); {access None}
   M352_M1_DR_IN_MAS : MOTION_INSTRUCTION := (FLAGS := -1442840576, EN := 1, DN := 1, PC := 1); {access None}
   M352_M1_DR_IN_MCD : MOTION_INSTRUCTION := (FLAGS := 570425344, DN := 1); {access None}
   M352_M1_DR_IN_MRP : MOTION_INSTRUCTION := (FLAGS := 33554432); {access None}
   M352_M1_DR_MAFR : MOTION_INSTRUCTION := (FLAGS := 301989888, ER := 1, ERR := 11); {access None}
   M352_M1_DR_MDR : MOTION_INSTRUCTION := (FLAGS := -1845493760, EN := 1, ER := 1, ERR := 11); {access None}
   M352_M1_DR_MSF : MOTION_INSTRUCTION := (FLAGS := 536870912, DN := 1, STATUS := 2, STATE := 1); {access None}
   M352_M1_DR_MSO : MOTION_INSTRUCTION := (FLAGS := -1577058304, EN := 1, DN := 1, STATE := 1); {access None}
   M352_M1_DR_OUT_MAJ : MOTION_INSTRUCTION := (FLAGS := 570425344, DN := 1); {access None}
   M352_M1_DR_OUT_MAM : MOTION_INSTRUCTION := (FLAGS := 33554432); {access None}
   M352_M1_DR_OUT_MAR : MOTION_INSTRUCTION := (FLAGS := 33554432); {access None}
   M352_M1_DR_OUT_MAS : MOTION_INSTRUCTION := (FLAGS := -1442840576, EN := 1, DN := 1, PC := 1); {access None}
   M352_M1_DR_OUT_MCD : MOTION_INSTRUCTION := (FLAGS := 570425344, DN := 1); {access None}
   M352_M1_DR_OUT_MRP : MOTION_INSTRUCTION := (FLAGS := 33554432); {access None}
   M352_ONS1 : BOOL;
   M352_ONS_SetResetPresence : BOOL;
   M352_Output_xAutoMode : BOOL := 1;
   M352_Output_xDescentBlockGlass : BOOL := 1;
   M352_Output_xGlassPresence : BOOL;
   M352_Output_xHA_Alarm : BOOL;   // W254HA1. Acustic alarm
   M352_Output_xHL_Alarm : BOOL;
   M352_Output_xHLReqGlass : BOOL;   // W204SB1. Glass sheet request
   M352_Output_xHLSendToCullet : BOOL;   // W204SB2. Sent to cullet
   M352_Output_xRiseBlockGlass : BOOL;
   M352_SpaceConv_Utilities : SpaceConv_Utilities := (CONST_dSyncMode := 1, CONST_dSyncroPhWindow_cmm := 200000, CONST_dConveyorLength_cmm := 500000, CONST_dConveyorWidth_cmm := 400000, CONST_dPresetFeedbackTime_ms := 500, CONST_rAcceleration_ms2 := 1.2, CONST_rDeceleration_ms2 := 1.2, CONF_MD1_dScan_ms := 20, CONF_MD4_MD6_dLength_cmm := 360000, CONF_MD7_dOffset_cmm := 50000, ST_xLastModLoadBkw := 1, ST_dStopLoadForseen_cmm := 495370, ST_dRealSpeed_mm_min := 40000, ST_rStepAdvancementH := 1333.3334, ST_rStepAdvancementT := 1333.3334, O_xPlateSynchronized := 1, O_dCountFeedbackTime_ms := 500, O_dPresetLoadUnload_cmm := -440770);
   M353 : MAC_Conveyor;
        .INPUT_xMotorThermalProbe_M1   // M315A.M1.Q403BT3. Motor thermal probe
        .PH_x.0   // Load
        .PH_x.1   // Load Upstream
        .PH_x.10   // Unload Downstream
        .PH_x.13   // End unload Upstream
        .PH_x.14   // End unload Downstream
        .PH_x.15   // End unload
        .PH_x.16   // Unpack convoy
        .PH_x.17   // End unpack convoy
        .PH_x.18   // Unpack convoy Upstream
        .PH_x.19   // End unpack convoy Upstream
        .PH_x.2   // Load Downstream
        .PH_x.20   // Unpack convoy Downstream
        .PH_x.21   // End unpack convoy Downstream
        .PH_x.22   // Stop for unload on main line
        .PH_x.23   // End stop for unload on main line
        .PH_x.24   // Stop for unload on main line Upstream
        .PH_x.25   // End stop for unload on main line Upstream
        .PH_x.26   // Stop for unload on main line Downstream
        .PH_x.27   // End stop for unload on main line Downstream
        .PH_x.28   // Load reentry
        .PH_x.29   // End load reentry
        .PH_x.5   // End load Upstream
        .PH_x.6   // End load Downstream
        .PH_x.7   // End load
        .PH_x.8   // Unload
        .PH_x.9   // Unload Upstream
   M353_ALM : MAC_Conveyor_ALM;
        .rgxWarning[0].0   // Z402.M315A.Q115B1.Plate not synchronized
        .rgxWarning[0].1   // Z402.M315A.Positioning error
   M353_Data : UDT_Convoy_SL;
   M353_HMR : MAC_Conveyor_HMR := (xManualCommandEnabled := 1, dState4 := 1);
        .dErrorCode1   // Error code M1
        .rgxMan.0   // Run M1
        .rgxMan.1   // Reverse M1
        .rgxMan.2   // Run M2
        .rgxMan.3   // Reverse M2
        .rgxMan.4   // Run M3
        .rgxMan.5   // Reverse M3
        .dErrorCode2   // Error code M2 (NU)
        .dErrorCode3   // Error code M3 (NU)
   M353_HMW : MAC_Conveyor_HMW;
        .rgxMan.0   // Run M1
        .rgxMan.1   // Reverse M1
        .rgxMan.2   // Run M2
        .rgxMan.3   // Reverse M2
        .rgxMan.4   // Run M3
        .rgxMan.5   // Reverse M3
   M353_M1_DR : AXIS_CIP_DRIVE; {access Read Only}
   M353_M1_DR_IN_MAJ : MOTION_INSTRUCTION := (FLAGS := 570425344, DN := 1); {access None}
   M353_M1_DR_IN_MAM : MOTION_INSTRUCTION := (FLAGS := 33554432); {access None}
   M353_M1_DR_IN_MAR : MOTION_INSTRUCTION := (FLAGS := 33554432); {access None}
   M353_M1_DR_IN_MAS : MOTION_INSTRUCTION := (FLAGS := -1442840576, EN := 1, DN := 1, PC := 1); {access None}
   M353_M1_DR_IN_MCD : MOTION_INSTRUCTION := (FLAGS := 570425344, DN := 1); {access None}
   M353_M1_DR_IN_MRP : MOTION_INSTRUCTION := (FLAGS := 33554432); {access None}
   M353_M1_DR_MAFR : MOTION_INSTRUCTION := (FLAGS := 301989888, ER := 1, ERR := 11); {access None}
   M353_M1_DR_MDR : MOTION_INSTRUCTION := (FLAGS := -1845493760, EN := 1, ER := 1, ERR := 11); {access None}
   M353_M1_DR_MSF : MOTION_INSTRUCTION := (FLAGS := 536870912, DN := 1, STATUS := 2, STATE := 1); {access None}
   M353_M1_DR_MSO : MOTION_INSTRUCTION := (FLAGS := -1577058304, EN := 1, DN := 1, STATE := 1); {access None}
   M353_M1_DR_OUT_MAJ : MOTION_INSTRUCTION := (FLAGS := 570425344, DN := 1); {access None}
   M353_M1_DR_OUT_MAM : MOTION_INSTRUCTION := (FLAGS := 33554432); {access None}
   M353_M1_DR_OUT_MAR : MOTION_INSTRUCTION := (FLAGS := 33554432); {access None}
   M353_M1_DR_OUT_MAS : MOTION_INSTRUCTION := (FLAGS := -1442840576, EN := 1, DN := 1, PC := 1); {access None}
   M353_M1_DR_OUT_MCD : MOTION_INSTRUCTION := (FLAGS := 570425344, DN := 1); {access None}
   M353_M1_DR_OUT_MRP : MOTION_INSTRUCTION := (FLAGS := 33554432); {access None}
   M353_SpaceConv_Utilities : SpaceConv_Utilities := (CONST_dSyncMode := 1, CONST_dSyncroPhWindow_cmm := 200000, CONST_dConveyorLength_cmm := 500000, CONST_dConveyorWidth_cmm := 400000, CONST_dPresetFeedbackTime_ms := 500, CONST_rAcceleration_ms2 := 1.2, CONST_rDeceleration_ms2 := 1.2, CONF_MD1_dScan_ms := 20, CONF_MD4_MD6_dLength_cmm := 360000, CONF_MD7_dOffset_cmm := 50000, ST_xLastModLoadBkw := 1, ST_dStopLoadForseen_cmm := 495370, ST_dRealSpeed_mm_min := 40000, ST_rStepAdvancementH := 1333.3334, ST_rStepAdvancementT := 1333.3334, O_xPlateSynchronized := 1, O_dCountFeedbackTime_ms := 500, O_dPresetLoadUnload_cmm := -440770);
   M360_M1_DR : AXIS_CIP_DRIVE; {access Read Only}
   M410_DATA_xSendERR : BOOL; {access Read Only}
   M420_DATA_xSendERR : BOOL;
   MCC1300_rgtDiagModule_HMI : GP_NetworkDiag_v1[90] := ([0].xConnected := 1, [0].dEntryStatus := 16#0000_4000, [0].dInstance := 16#0000_0a6d, [1].xConnected := 1, [1].dEntryStatus := 16#0000_4000, [1].dInstance := 16#0000_095f, [2].xConnected := 1, [2].dEntryStatus := 16#0000_4000, [2].dInstance := 16#0000_a3f5, [3].xConnected := 1, [3].dEntryStatus := 16#0000_4000, [3].dInstance := 16#0000_ba43, [4].xConnected := 1, [4].dEntryStatus := 16#0000_4000, [4].dInstance := 16#0000_af16, [5].xConnected := 1, [5].dEntryStatus := 16#0000_4000, [5].dInstance := 16#0000_5f5d, [9].xConnected := 1, [9].dEntryStatus := 16#0000_4000, [9].dInstance := 16#0000_3ec5, [10].xConnected := 1, [10].dEntryStatus := 16#0000_4000, [10].dInstance := 16#0000_5f5d, [11].xConnected := 1, [11].dEntryStatus := 16#0000_4000, [11].dInstance := 16#0000_6b09, [12].xConnected := 1, [12].dEntryStatus := 16#0000_4000, [12].dInstance := 16#0000_6808, [13].xConnected := 1, [13].dEntryStatus := 16#0000_4000, [13].dInstance := 16#0000_ba5f, [14].xConnected := 1, [14].dEntryStatus := 16#0000_4000, [14].dInstance := 16#0000_c7c6, [15].xConnected := 1, [15].dEntryStatus := 16#0000_4000, [15].dInstance := 16#0000_0bf1, [16].xConnected := 1, [16].dEntryStatus := 16#0000_4000, [16].dInstance := 16#0000_3650, [17].xConnected := 1, [17].dEntryStatus := 16#0000_4000, [17].dInstance := 16#0000_9e93, [18].xConnected := 1, [18].dEntryStatus := 16#0000_4000, [18].dInstance := 16#0000_cbaa, [19].xConnected := 1, [19].dEntryStatus := 16#0000_4000, [19].dInstance := 16#0000_7c6b, [20].xConnected := 1, [20].dEntryStatus := 16#0000_4000, [20].dInstance := 16#0000_b922, [21].xConnected := 1, [21].dEntryStatus := 16#0000_4000, [21].dInstance := 16#0000_415d, [22].xConnected := 1, [22].dEntryStatus := 16#0000_4000, [22].dInstance := 16#0000_698c,
        [23].xConnected := 1, [23].dEntryStatus := 16#0000_4000, [23].dInstance := 16#0000_f254, [24].xConnected := 1, [24].xFaulted := 1, [24].dEntryStatus := 16#0000_3000, [24].dFaultCode := 16#0000_0204, [24].dInstance := 16#0000_1662, [25].xFaulted := 1, [25].dEntryStatus := 16#0000_1000, [25].dFaultCode := 16#0000_0204, [25].dInstance := 16#0000_719d, [26].xConnected := 1, [26].xFaulted := 1, [26].dEntryStatus := 16#0000_3000, [26].dFaultCode := 16#0000_0204, [26].dInstance := 16#0000_00cc, [27].xFaulted := 1, [27].dEntryStatus := 16#0000_1000, [27].dFaultCode := 16#0000_0204, [27].dInstance := 16#0000_7c9f, [28].xConnected := 1, [28].xFaulted := 1, [28].dEntryStatus := 16#0000_3000, [28].dFaultCode := 16#0000_0204, [28].dInstance := 16#0000_e906, [29].xConnected := 1, [29].xFaulted := 1, [29].dEntryStatus := 16#0000_3000, [29].dFaultCode := 16#0000_0204, [29].dInstance := 16#0000_7031, [30].xConnected := 1, [30].xFaulted := 1, [30].dEntryStatus := 16#0000_3000, [30].dFaultCode := 16#0000_0204, [30].dInstance := 16#0000_cda9, [31].xConnected := 1, [31].xFaulted := 1, [31].dEntryStatus := 16#0000_3000, [31].dFaultCode := 16#0000_0204, [31].dInstance := 16#0000_b190, [32].xFaulted := 1, [32].dEntryStatus := 16#0000_1000, [32].dFaultCode := 16#0000_0204, [32].dInstance := 16#0000_7a24, [33].xConnected := 1, [33].xFaulted := 1, [33].dEntryStatus := 16#0000_3000, [33].dFaultCode := 16#0000_0204, [33].dInstance := 16#0000_c797, [34].xConnected := 1, [34].xFaulted := 1, [34].dEntryStatus := 16#0000_3000, [34].dFaultCode := 16#0000_0204, [34].dInstance := 16#0000_431e, [35].xFaulted := 1, [35].dEntryStatus := 16#0000_1000, [35].dFaultCode := 16#0000_0204, [35].dInstance := 16#0000_90e9, [36].xConnected := 1,
